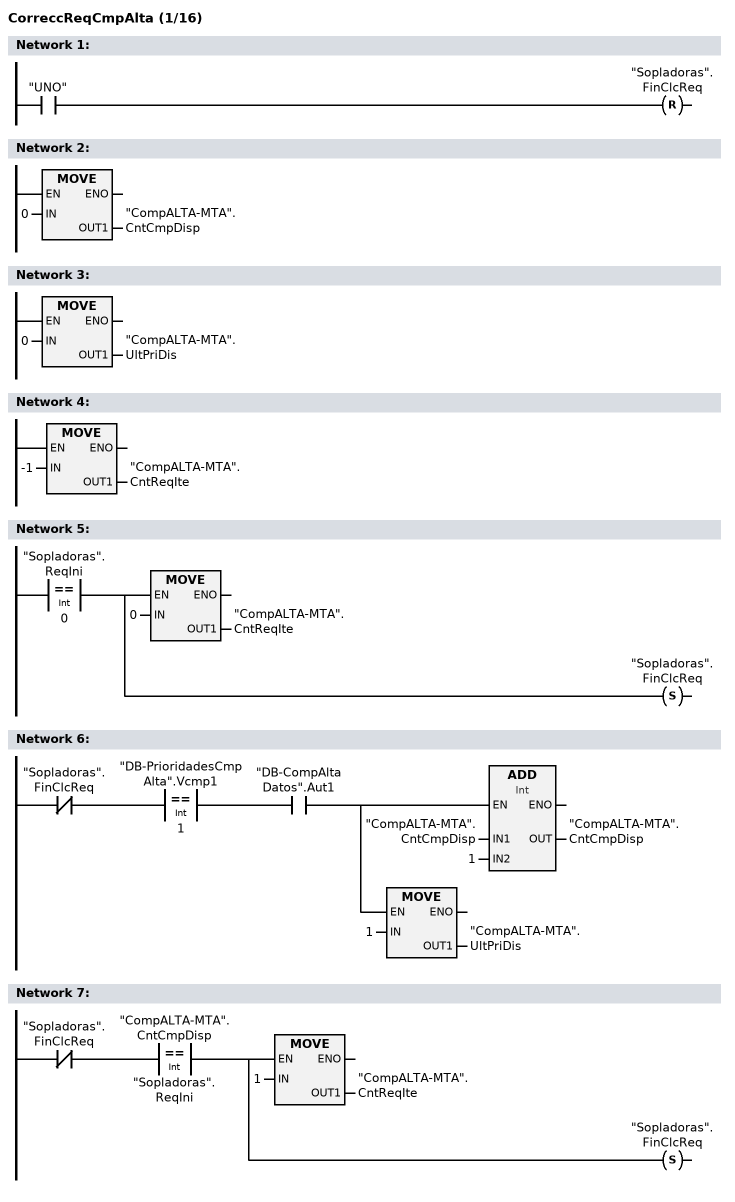
   RUNG wire#powerrail
      Contact( "UNO" )
      R_Coil( "Sopladoras".FinClcReq )
   END_RUNG
   // the same network as SCL:
   IF "UNO" THEN "Sopladoras".FinClcReq := FALSE; END_IF;
END_REGION

REGION Network 2
   RUNG wire#powerrail
      { S7_GenerateENO := "TRUE" } Move(in := 0, out1 => "CompALTA-MTA".CntCmpDisp)
   END_RUNG
   // the same network as SCL:
   "CompALTA-MTA".CntCmpDisp := 0;
END_REGION

REGION Network 3
   RUNG wire#powerrail
      { S7_GenerateENO := "TRUE" } Move(in := 0, out1 => "CompALTA-MTA".UltPriDis)
   END_RUNG
   // the same network as SCL:
   "CompALTA-MTA".UltPriDis := 0;
END_REGION

REGION Network 4
   RUNG wire#powerrail
      { S7_GenerateENO := "TRUE" } Move(in := -1, out1 => "CompALTA-MTA".CntReqIte)
   END_RUNG
   // the same network as SCL:
   "CompALTA-MTA".CntReqIte := -1;
END_REGION

REGION Network 5
   RUNG wire#powerrail
      { S7_Templates := "SrcType := Int" } EQ_Contact(in1 := "Sopladoras".ReqIni, in2 := 0)
      wire#w1
      { S7_GenerateENO := "TRUE" } Move(in := 0, out1 => "CompALTA-MTA".CntReqIte)
   END_RUNG
   RUNG wire#w1
      S_Coil( "Sopladoras".FinClcReq )
   END_RUNG
   // the same network as SCL:
   IF "Sopladoras".ReqIni = 0 THEN
       "CompALTA-MTA".CntReqIte := 0;
       "Sopladoras".FinClcReq := TRUE;
   END_IF;
END_REGION

REGION Network 6
   IF NOT "Sopladoras".FinClcReq AND ("DB-PrioridadesCmpAlta".Vcmp1 = 1) AND "DB-CompAltaDatos".Aut1 THEN
       "CompALTA-MTA".CntCmpDisp := "CompALTA-MTA".CntCmpDisp + 1;
       "CompALTA-MTA".UltPriDis := 1;
   END_IF;
END_REGION

REGION Network 7
   IF NOT "Sopladoras".FinClcReq AND ("CompALTA-MTA".CntCmpDisp = "Sopladoras".ReqIni) THEN
       "CompALTA-MTA".CntReqIte := 1;
       "Sopladoras".FinClcReq := TRUE;
   END_IF;
END_REGION

REGION Network 8
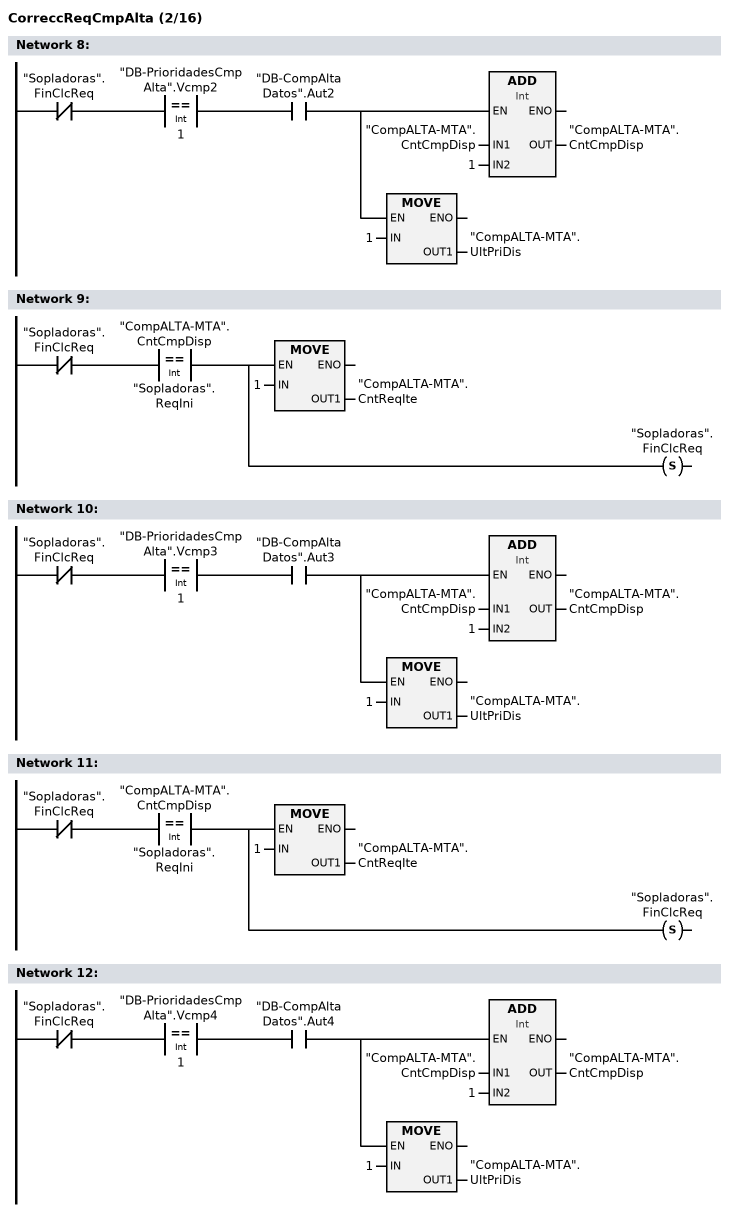
   IF NOT "Sopladoras".FinClcReq AND ("DB-PrioridadesCmpAlta".Vcmp2 = 1) AND "DB-CompAltaDatos".Aut2 THEN
       "CompALTA-MTA".CntCmpDisp := "CompALTA-MTA".CntCmpDisp + 1;
       "CompALTA-MTA".UltPriDis := 1;
   END_IF;
END_REGION

REGION Network 9
   IF NOT "Sopladoras".FinClcReq AND ("CompALTA-MTA".CntCmpDisp = "Sopladoras".ReqIni) THEN
       "CompALTA-MTA".CntReqIte := 1;
       "Sopladoras".FinClcReq := TRUE;
   END_IF;
END_REGION

REGION Network 10
   IF NOT "Sopladoras".FinClcReq AND ("DB-PrioridadesCmpAlta".Vcmp3 = 1) AND "DB-CompAltaDatos".Aut3 THEN
       "CompALTA-MTA".CntCmpDisp := "CompALTA-MTA".CntCmpDisp + 1;
       "CompALTA-MTA".UltPriDis := 1;
   END_IF;
END_REGION

REGION Network 11
   IF NOT "Sopladoras".FinClcReq AND ("CompALTA-MTA".CntCmpDisp = "Sopladoras".ReqIni) THEN
       "CompALTA-MTA".CntReqIte := 1;
       "Sopladoras".FinClcReq := TRUE;
   END_IF;
END_REGION

REGION Network 12
   IF NOT "Sopladoras".FinClcReq AND ("DB-PrioridadesCmpAlta".Vcmp4 = 1) AND "DB-CompAltaDatos".Aut4 THEN
       "CompALTA-MTA".CntCmpDisp := "CompALTA-MTA".CntCmpDisp + 1;
       "CompALTA-MTA".UltPriDis := 1;
   END_IF;
END_REGION

REGION Network 13
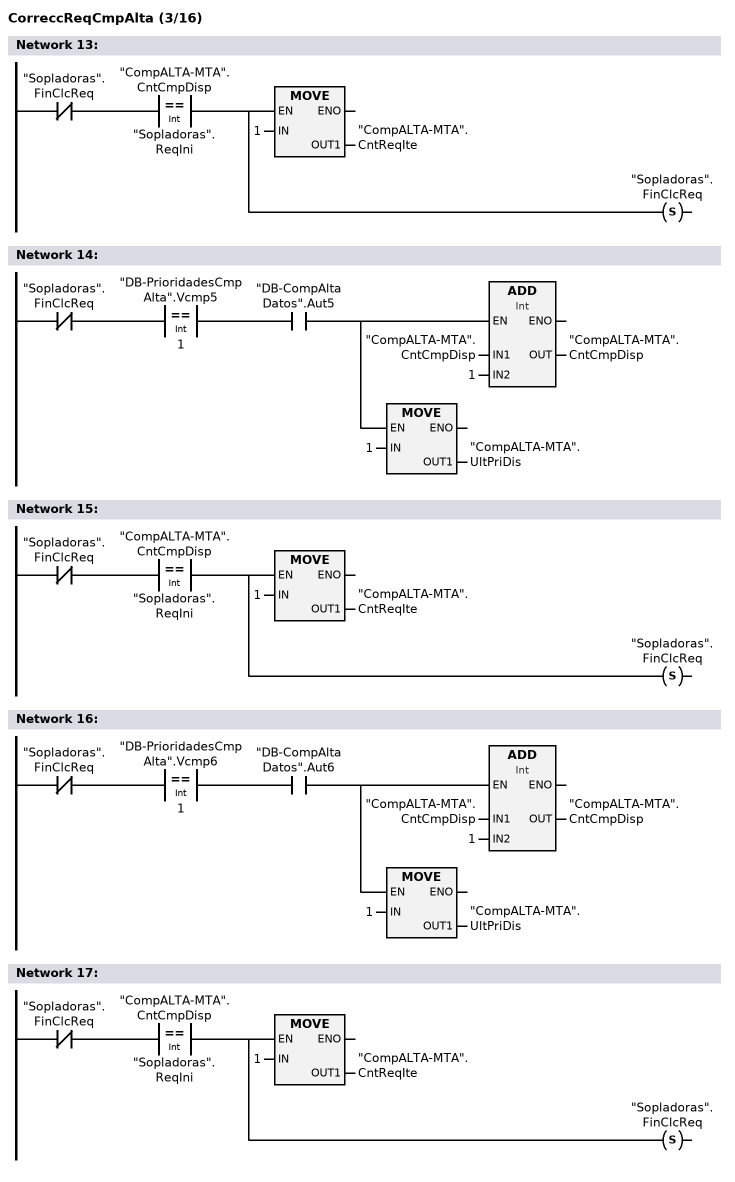
   IF NOT "Sopladoras".FinClcReq AND ("CompALTA-MTA".CntCmpDisp = "Sopladoras".ReqIni) THEN
       "CompALTA-MTA".CntReqIte := 1;
       "Sopladoras".FinClcReq := TRUE;
   END_IF;
END_REGION

REGION Network 14
   IF NOT "Sopladoras".FinClcReq AND ("DB-PrioridadesCmpAlta".Vcmp5 = 1) AND "DB-CompAltaDatos".Aut5 THEN
       "CompALTA-MTA".CntCmpDisp := "CompALTA-MTA".CntCmpDisp + 1;
       "CompALTA-MTA".UltPriDis := 1;
   END_IF;
END_REGION

REGION Network 15
   IF NOT "Sopladoras".FinClcReq AND ("CompALTA-MTA".CntCmpDisp = "Sopladoras".ReqIni) THEN
       "CompALTA-MTA".CntReqIte := 1;
       "Sopladoras".FinClcReq := TRUE;
   END_IF;
END_REGION

REGION Network 16
   RUNG wire#powerrail
      I_Contact( "Sopladoras".FinClcReq )
      { S7_Templates := "SrcType := Int" } EQ_Contact(in1 := "DB-PrioridadesCmpAlta".Vcmp6, in2 := 1)
      Contact( "DB-CompAltaDatos".Aut6 )
      wire#w1
      { S7_Templates := "SrcType := Int"; S7_GenerateENO := "TRUE" } Add(in1 := "CompALTA-MTA".CntCmpDisp, in2 := 1, out => "CompALTA-MTA".CntCmpDisp)
   END_RUNG
   RUNG wire#w1
      { S7_GenerateENO := "TRUE" } Move(in := 1, out1 => "CompALTA-MTA".UltPriDis)
   END_RUNG
   // the same network as SCL:
   IF NOT "Sopladoras".FinClcReq AND ("DB-PrioridadesCmpAlta".Vcmp6 = 1) AND "DB-CompAltaDatos".Aut6 THEN
       "CompALTA-MTA".CntCmpDisp := "CompALTA-MTA".CntCmpDisp + 1;
       "CompALTA-MTA".UltPriDis := 1;
   END_IF;
END_REGION

REGION Network 17
   RUNG wire#powerrail
      I_Contact( "Sopladoras".FinClcReq )
      { S7_Templates := "SrcType := Int" } EQ_Contact(in1 := "CompALTA-MTA".CntCmpDisp, in2 := "Sopladoras".ReqIni)
      wire#w1
      { S7_GenerateENO := "TRUE" } Move(in := 1, out1 => "CompALTA-MTA".CntReqIte)
   END_RUNG
   RUNG wire#w1
      S_Coil( "Sopladoras".FinClcReq )
   END_RUNG
   // the same network as SCL:
   IF NOT "Sopladoras".FinClcReq AND ("CompALTA-MTA".CntCmpDisp = "Sopladoras".ReqIni) THEN
       "CompALTA-MTA".CntReqIte := 1;
       "Sopladoras".FinClcReq := TRUE;
   END_IF;
END_REGION

REGION Network 18
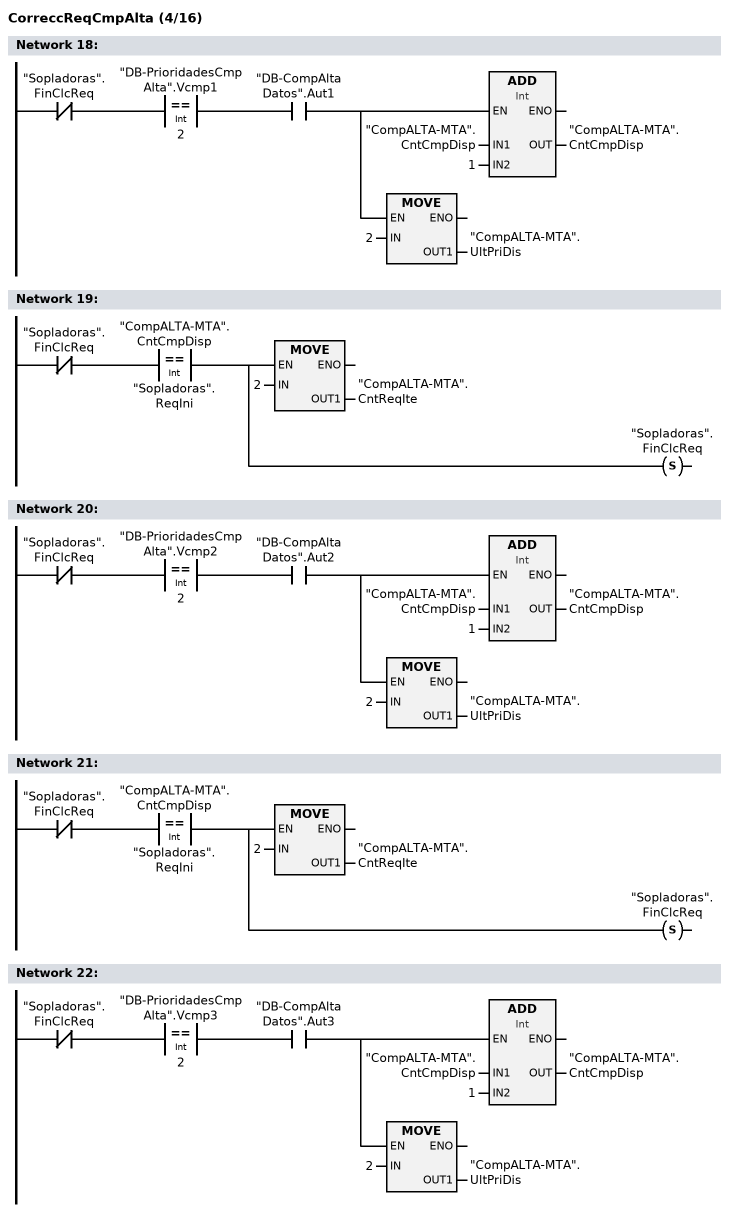
   IF NOT "Sopladoras".FinClcReq AND ("DB-PrioridadesCmpAlta".Vcmp1 = 2) AND "DB-CompAltaDatos".Aut1 THEN
       "CompALTA-MTA".CntCmpDisp := "CompALTA-MTA".CntCmpDisp + 1;
       "CompALTA-MTA".UltPriDis := 2;
   END_IF;
END_REGION

REGION Network 19
   IF NOT "Sopladoras".FinClcReq AND ("CompALTA-MTA".CntCmpDisp = "Sopladoras".ReqIni) THEN
       "CompALTA-MTA".CntReqIte := 2;
       "Sopladoras".FinClcReq := TRUE;
   END_IF;
END_REGION

REGION Network 20
   IF NOT "Sopladoras".FinClcReq AND ("DB-PrioridadesCmpAlta".Vcmp2 = 2) AND "DB-CompAltaDatos".Aut2 THEN
       "CompALTA-MTA".CntCmpDisp := "CompALTA-MTA".CntCmpDisp + 1;
       "CompALTA-MTA".UltPriDis := 2;
   END_IF;
END_REGION

REGION Network 21
   IF NOT "Sopladoras".FinClcReq AND ("CompALTA-MTA".CntCmpDisp = "Sopladoras".ReqIni) THEN
       "CompALTA-MTA".CntReqIte := 2;
       "Sopladoras".FinClcReq := TRUE;
   END_IF;
END_REGION

REGION Network 22
   IF NOT "Sopladoras".FinClcReq AND ("DB-PrioridadesCmpAlta".Vcmp3 = 2) AND "DB-CompAltaDatos".Aut3 THEN
       "CompALTA-MTA".CntCmpDisp := "CompALTA-MTA".CntCmpDisp + 1;
       "CompALTA-MTA".UltPriDis := 2;
   END_IF;
END_REGION

REGION Network 23
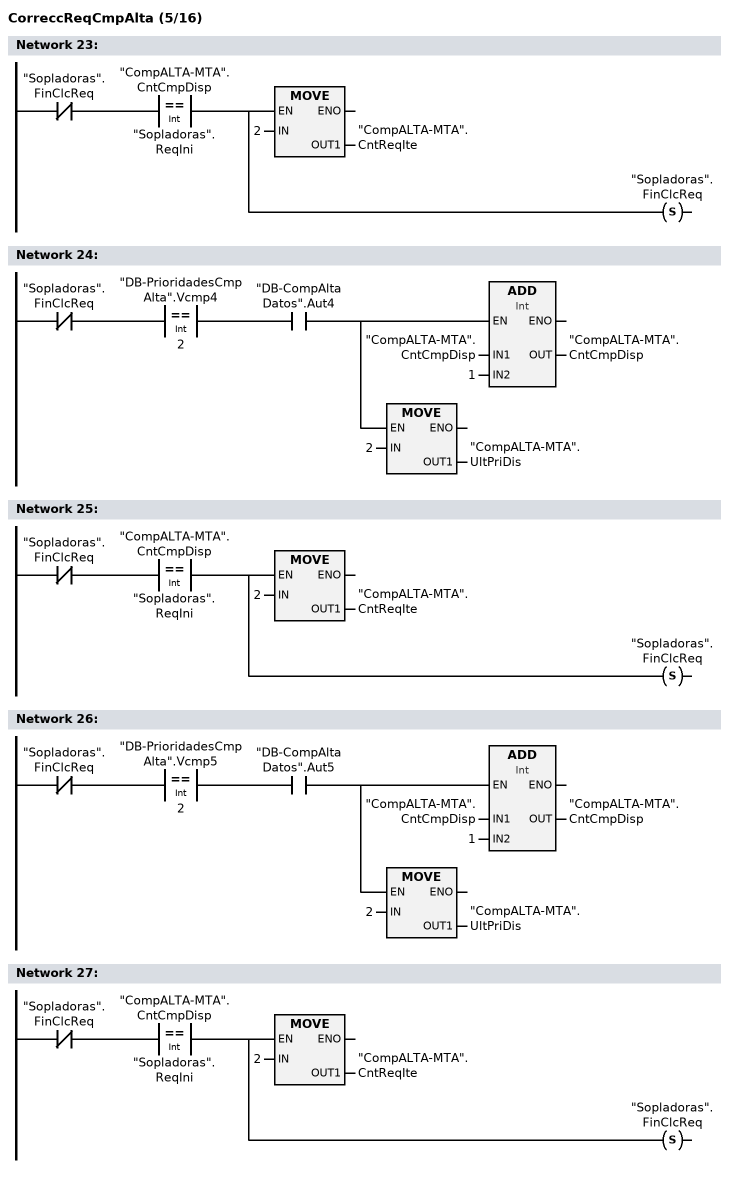
   IF NOT "Sopladoras".FinClcReq AND ("CompALTA-MTA".CntCmpDisp = "Sopladoras".ReqIni) THEN
       "CompALTA-MTA".CntReqIte := 2;
       "Sopladoras".FinClcReq := TRUE;
   END_IF;
END_REGION

REGION Network 24
   IF NOT "Sopladoras".FinClcReq AND ("DB-PrioridadesCmpAlta".Vcmp4 = 2) AND "DB-CompAltaDatos".Aut4 THEN
       "CompALTA-MTA".CntCmpDisp := "CompALTA-MTA".CntCmpDisp + 1;
       "CompALTA-MTA".UltPriDis := 2;
   END_IF;
END_REGION

REGION Network 25
   IF NOT "Sopladoras".FinClcReq AND ("CompALTA-MTA".CntCmpDisp = "Sopladoras".ReqIni) THEN
       "CompALTA-MTA".CntReqIte := 2;
       "Sopladoras".FinClcReq := TRUE;
   END_IF;
END_REGION

REGION Network 26
   IF NOT "Sopladoras".FinClcReq AND ("DB-PrioridadesCmpAlta".Vcmp5 = 2) AND "DB-CompAltaDatos".Aut5 THEN
       "CompALTA-MTA".CntCmpDisp := "CompALTA-MTA".CntCmpDisp + 1;
       "CompALTA-MTA".UltPriDis := 2;
   END_IF;
END_REGION

REGION Network 27
   IF NOT "Sopladoras".FinClcReq AND ("CompALTA-MTA".CntCmpDisp = "Sopladoras".ReqIni) THEN
       "CompALTA-MTA".CntReqIte := 2;
       "Sopladoras".FinClcReq := TRUE;
   END_IF;
END_REGION

REGION Network 28
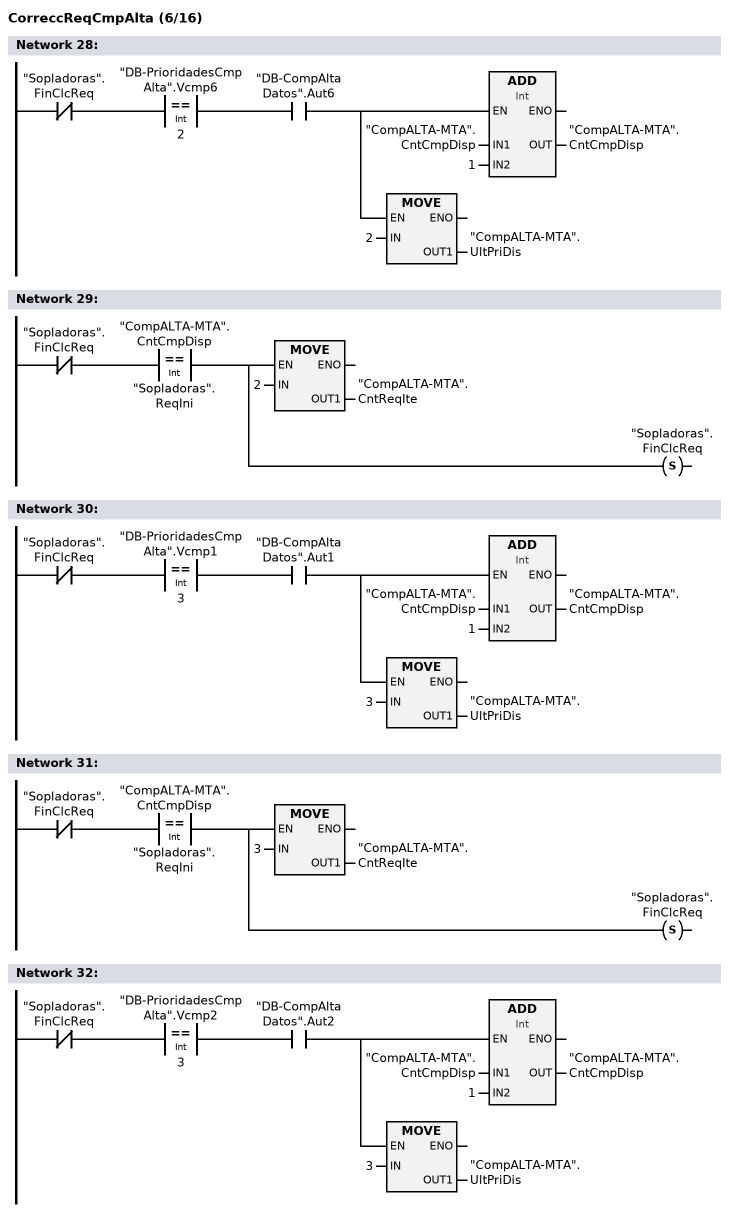
   RUNG wire#powerrail
      I_Contact( "Sopladoras".FinClcReq )
      { S7_Templates := "SrcType := Int" } EQ_Contact(in1 := "DB-PrioridadesCmpAlta".Vcmp6, in2 := 2)
      Contact( "DB-CompAltaDatos".Aut6 )
      wire#w1
      { S7_Templates := "SrcType := Int"; S7_GenerateENO := "TRUE" } Add(in1 := "CompALTA-MTA".CntCmpDisp, in2 := 1, out => "CompALTA-MTA".CntCmpDisp)
   END_RUNG
   RUNG wire#w1
      { S7_GenerateENO := "TRUE" } Move(in := 2, out1 => "CompALTA-MTA".UltPriDis)
   END_RUNG
   // the same network as SCL:
   IF NOT "Sopladoras".FinClcReq AND ("DB-PrioridadesCmpAlta".Vcmp6 = 2) AND "DB-CompAltaDatos".Aut6 THEN
       "CompALTA-MTA".CntCmpDisp := "CompALTA-MTA".CntCmpDisp + 1;
       "CompALTA-MTA".UltPriDis := 2;
   END_IF;
END_REGION

REGION Network 29
   RUNG wire#powerrail
      I_Contact( "Sopladoras".FinClcReq )
      { S7_Templates := "SrcType := Int" } EQ_Contact(in1 := "CompALTA-MTA".CntCmpDisp, in2 := "Sopladoras".ReqIni)
      wire#w1
      { S7_GenerateENO := "TRUE" } Move(in := 2, out1 => "CompALTA-MTA".CntReqIte)
   END_RUNG
   RUNG wire#w1
      S_Coil( "Sopladoras".FinClcReq )
   END_RUNG
   // the same network as SCL:
   IF NOT "Sopladoras".FinClcReq AND ("CompALTA-MTA".CntCmpDisp = "Sopladoras".ReqIni) THEN
       "CompALTA-MTA".CntReqIte := 2;
       "Sopladoras".FinClcReq := TRUE;
   END_IF;
END_REGION

REGION Network 30
   IF NOT "Sopladoras".FinClcReq AND ("DB-PrioridadesCmpAlta".Vcmp1 = 3) AND "DB-CompAltaDatos".Aut1 THEN
       "CompALTA-MTA".CntCmpDisp := "CompALTA-MTA".CntCmpDisp + 1;
       "CompALTA-MTA".UltPriDis := 3;
   END_IF;
END_REGION

REGION Network 31
   IF NOT "Sopladoras".FinClcReq AND ("CompALTA-MTA".CntCmpDisp = "Sopladoras".ReqIni) THEN
       "CompALTA-MTA".CntReqIte := 3;
       "Sopladoras".FinClcReq := TRUE;
   END_IF;
END_REGION

REGION Network 32
   IF NOT "Sopladoras".FinClcReq AND ("DB-PrioridadesCmpAlta".Vcmp2 = 3) AND "DB-CompAltaDatos".Aut2 THEN
       "CompALTA-MTA".CntCmpDisp := "CompALTA-MTA".CntCmpDisp + 1;
       "CompALTA-MTA".UltPriDis := 3;
   END_IF;
END_REGION

REGION Network 33
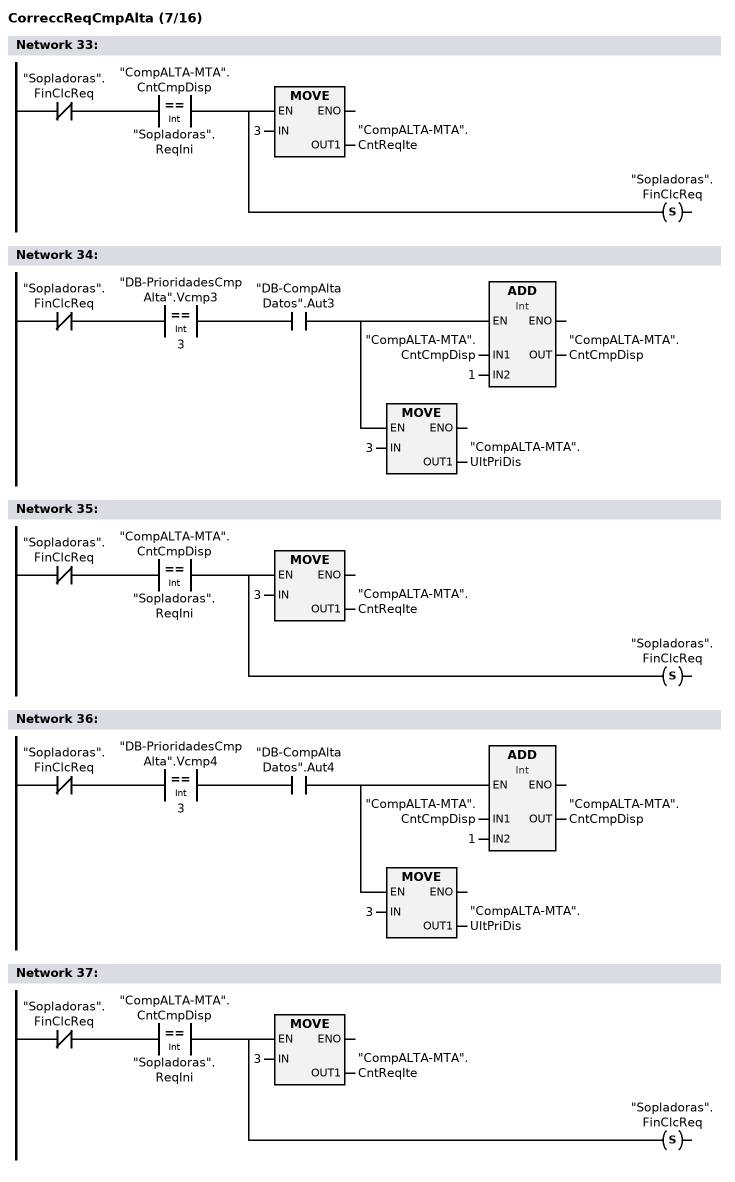
   IF NOT "Sopladoras".FinClcReq AND ("CompALTA-MTA".CntCmpDisp = "Sopladoras".ReqIni) THEN
       "CompALTA-MTA".CntReqIte := 3;
       "Sopladoras".FinClcReq := TRUE;
   END_IF;
END_REGION

REGION Network 34
   IF NOT "Sopladoras".FinClcReq AND ("DB-PrioridadesCmpAlta".Vcmp3 = 3) AND "DB-CompAltaDatos".Aut3 THEN
       "CompALTA-MTA".CntCmpDisp := "CompALTA-MTA".CntCmpDisp + 1;
       "CompALTA-MTA".UltPriDis := 3;
   END_IF;
END_REGION

REGION Network 35
   IF NOT "Sopladoras".FinClcReq AND ("CompALTA-MTA".CntCmpDisp = "Sopladoras".ReqIni) THEN
       "CompALTA-MTA".CntReqIte := 3;
       "Sopladoras".FinClcReq := TRUE;
   END_IF;
END_REGION

REGION Network 36
   IF NOT "Sopladoras".FinClcReq AND ("DB-PrioridadesCmpAlta".Vcmp4 = 3) AND "DB-CompAltaDatos".Aut4 THEN
       "CompALTA-MTA".CntCmpDisp := "CompALTA-MTA".CntCmpDisp + 1;
       "CompALTA-MTA".UltPriDis := 3;
   END_IF;
END_REGION

REGION Network 37
   IF NOT "Sopladoras".FinClcReq AND ("CompALTA-MTA".CntCmpDisp = "Sopladoras".ReqIni) THEN
       "CompALTA-MTA".CntReqIte := 3;
       "Sopladoras".FinClcReq := TRUE;
   END_IF;
END_REGION

REGION Network 38
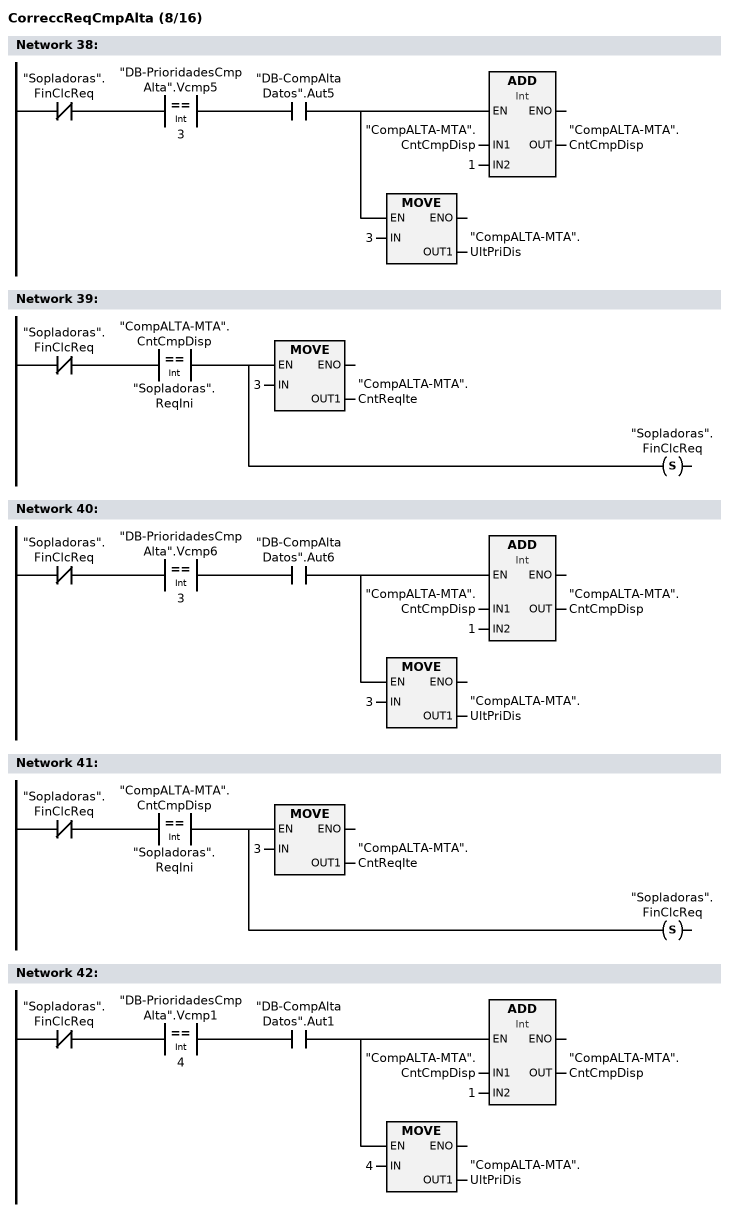
   IF NOT "Sopladoras".FinClcReq AND ("DB-PrioridadesCmpAlta".Vcmp5 = 3) AND "DB-CompAltaDatos".Aut5 THEN
       "CompALTA-MTA".CntCmpDisp := "CompALTA-MTA".CntCmpDisp + 1;
       "CompALTA-MTA".UltPriDis := 3;
   END_IF;
END_REGION

REGION Network 39
   IF NOT "Sopladoras".FinClcReq AND ("CompALTA-MTA".CntCmpDisp = "Sopladoras".ReqIni) THEN
       "CompALTA-MTA".CntReqIte := 3;
       "Sopladoras".FinClcReq := TRUE;
   END_IF;
END_REGION

REGION Network 40
   RUNG wire#powerrail
      I_Contact( "Sopladoras".FinClcReq )
      { S7_Templates := "SrcType := Int" } EQ_Contact(in1 := "DB-PrioridadesCmpAlta".Vcmp6, in2 := 3)
      Contact( "DB-CompAltaDatos".Aut6 )
      wire#w1
      { S7_Templates := "SrcType := Int"; S7_GenerateENO := "TRUE" } Add(in1 := "CompALTA-MTA".CntCmpDisp, in2 := 1, out => "CompALTA-MTA".CntCmpDisp)
   END_RUNG
   RUNG wire#w1
      { S7_GenerateENO := "TRUE" } Move(in := 3, out1 => "CompALTA-MTA".UltPriDis)
   END_RUNG
   // the same network as SCL:
   IF NOT "Sopladoras".FinClcReq AND ("DB-PrioridadesCmpAlta".Vcmp6 = 3) AND "DB-CompAltaDatos".Aut6 THEN
       "CompALTA-MTA".CntCmpDisp := "CompALTA-MTA".CntCmpDisp + 1;
       "CompALTA-MTA".UltPriDis := 3;
   END_IF;
END_REGION

REGION Network 41
   RUNG wire#powerrail
      I_Contact( "Sopladoras".FinClcReq )
      { S7_Templates := "SrcType := Int" } EQ_Contact(in1 := "CompALTA-MTA".CntCmpDisp, in2 := "Sopladoras".ReqIni)
      wire#w1
      { S7_GenerateENO := "TRUE" } Move(in := 3, out1 => "CompALTA-MTA".CntReqIte)
   END_RUNG
   RUNG wire#w1
      S_Coil( "Sopladoras".FinClcReq )
   END_RUNG
   // the same network as SCL:
   IF NOT "Sopladoras".FinClcReq AND ("CompALTA-MTA".CntCmpDisp = "Sopladoras".ReqIni) THEN
       "CompALTA-MTA".CntReqIte := 3;
       "Sopladoras".FinClcReq := TRUE;
   END_IF;
END_REGION

REGION Network 42
   IF NOT "Sopladoras".FinClcReq AND ("DB-PrioridadesCmpAlta".Vcmp1 = 4) AND "DB-CompAltaDatos".Aut1 THEN
       "CompALTA-MTA".CntCmpDisp := "CompALTA-MTA".CntCmpDisp + 1;
       "CompALTA-MTA".UltPriDis := 4;
   END_IF;
END_REGION

REGION Network 43
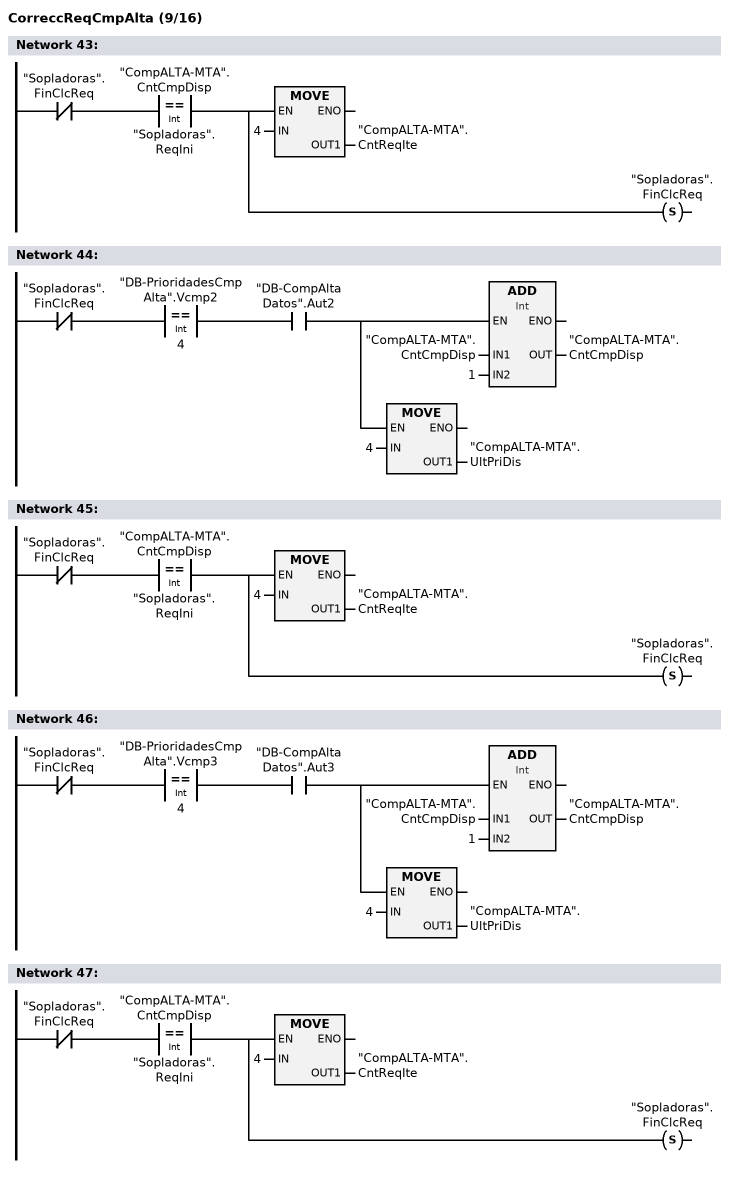
   IF NOT "Sopladoras".FinClcReq AND ("CompALTA-MTA".CntCmpDisp = "Sopladoras".ReqIni) THEN
       "CompALTA-MTA".CntReqIte := 4;
       "Sopladoras".FinClcReq := TRUE;
   END_IF;
END_REGION

REGION Network 44
   IF NOT "Sopladoras".FinClcReq AND ("DB-PrioridadesCmpAlta".Vcmp2 = 4) AND "DB-CompAltaDatos".Aut2 THEN
       "CompALTA-MTA".CntCmpDisp := "CompALTA-MTA".CntCmpDisp + 1;
       "CompALTA-MTA".UltPriDis := 4;
   END_IF;
END_REGION

REGION Network 45
   IF NOT "Sopladoras".FinClcReq AND ("CompALTA-MTA".CntCmpDisp = "Sopladoras".ReqIni) THEN
       "CompALTA-MTA".CntReqIte := 4;
       "Sopladoras".FinClcReq := TRUE;
   END_IF;
END_REGION

REGION Network 46
   IF NOT "Sopladoras".FinClcReq AND ("DB-PrioridadesCmpAlta".Vcmp3 = 4) AND "DB-CompAltaDatos".Aut3 THEN
       "CompALTA-MTA".CntCmpDisp := "CompALTA-MTA".CntCmpDisp + 1;
       "CompALTA-MTA".UltPriDis := 4;
   END_IF;
END_REGION

REGION Network 47
   IF NOT "Sopladoras".FinClcReq AND ("CompALTA-MTA".CntCmpDisp = "Sopladoras".ReqIni) THEN
       "CompALTA-MTA".CntReqIte := 4;
       "Sopladoras".FinClcReq := TRUE;
   END_IF;
END_REGION

REGION Network 48
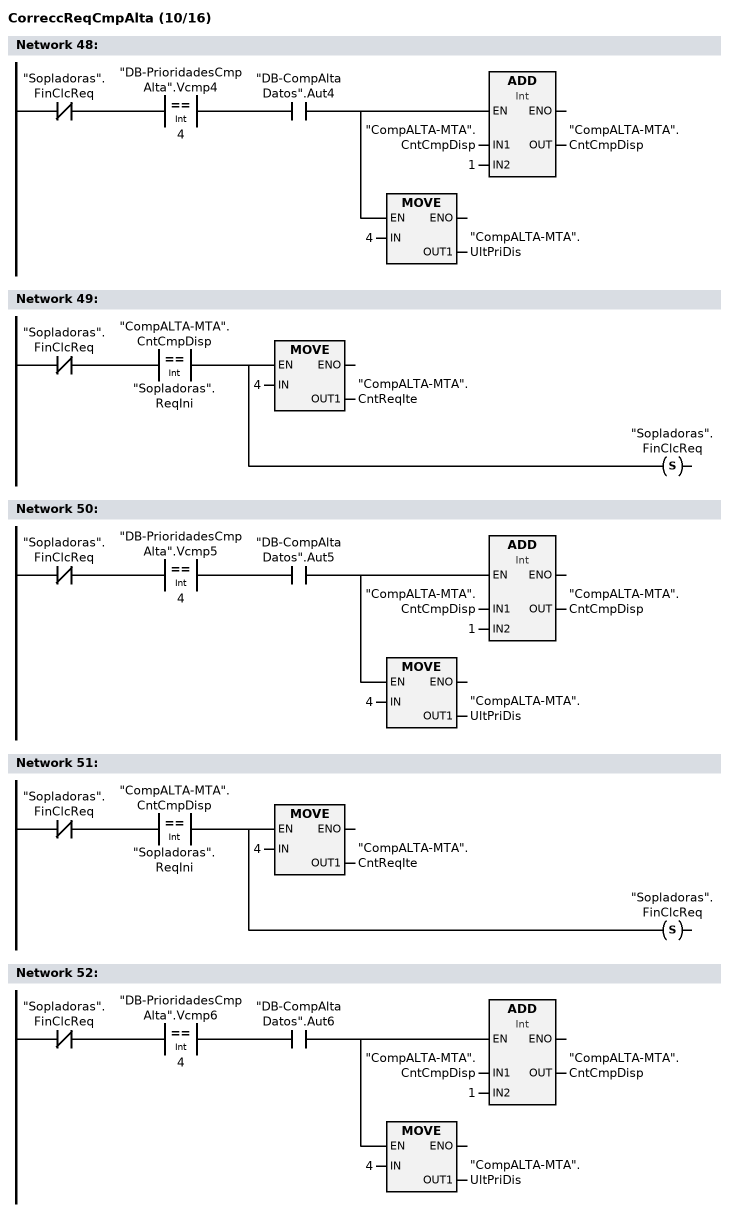
   IF NOT "Sopladoras".FinClcReq AND ("DB-PrioridadesCmpAlta".Vcmp4 = 4) AND "DB-CompAltaDatos".Aut4 THEN
       "CompALTA-MTA".CntCmpDisp := "CompALTA-MTA".CntCmpDisp + 1;
       "CompALTA-MTA".UltPriDis := 4;
   END_IF;
END_REGION

REGION Network 49
   IF NOT "Sopladoras".FinClcReq AND ("CompALTA-MTA".CntCmpDisp = "Sopladoras".ReqIni) THEN
       "CompALTA-MTA".CntReqIte := 4;
       "Sopladoras".FinClcReq := TRUE;
   END_IF;
END_REGION

REGION Network 50
   IF NOT "Sopladoras".FinClcReq AND ("DB-PrioridadesCmpAlta".Vcmp5 = 4) AND "DB-CompAltaDatos".Aut5 THEN
       "CompALTA-MTA".CntCmpDisp := "CompALTA-MTA".CntCmpDisp + 1;
       "CompALTA-MTA".UltPriDis := 4;
   END_IF;
END_REGION

REGION Network 51
   IF NOT "Sopladoras".FinClcReq AND ("CompALTA-MTA".CntCmpDisp = "Sopladoras".ReqIni) THEN
       "CompALTA-MTA".CntReqIte := 4;
       "Sopladoras".FinClcReq := TRUE;
   END_IF;
END_REGION

REGION Network 52
   RUNG wire#powerrail
      I_Contact( "Sopladoras".FinClcReq )
      { S7_Templates := "SrcType := Int" } EQ_Contact(in1 := "DB-PrioridadesCmpAlta".Vcmp6, in2 := 4)
      Contact( "DB-CompAltaDatos".Aut6 )
      wire#w1
      { S7_Templates := "SrcType := Int"; S7_GenerateENO := "TRUE" } Add(in1 := "CompALTA-MTA".CntCmpDisp, in2 := 1, out => "CompALTA-MTA".CntCmpDisp)
   END_RUNG
   RUNG wire#w1
      { S7_GenerateENO := "TRUE" } Move(in := 4, out1 => "CompALTA-MTA".UltPriDis)
   END_RUNG
   // the same network as SCL:
   IF NOT "Sopladoras".FinClcReq AND ("DB-PrioridadesCmpAlta".Vcmp6 = 4) AND "DB-CompAltaDatos".Aut6 THEN
       "CompALTA-MTA".CntCmpDisp := "CompALTA-MTA".CntCmpDisp + 1;
       "CompALTA-MTA".UltPriDis := 4;
   END_IF;
END_REGION

REGION Network 53